// TIA Portal project "uppgift2IndustriellIT" (V18) (continued)
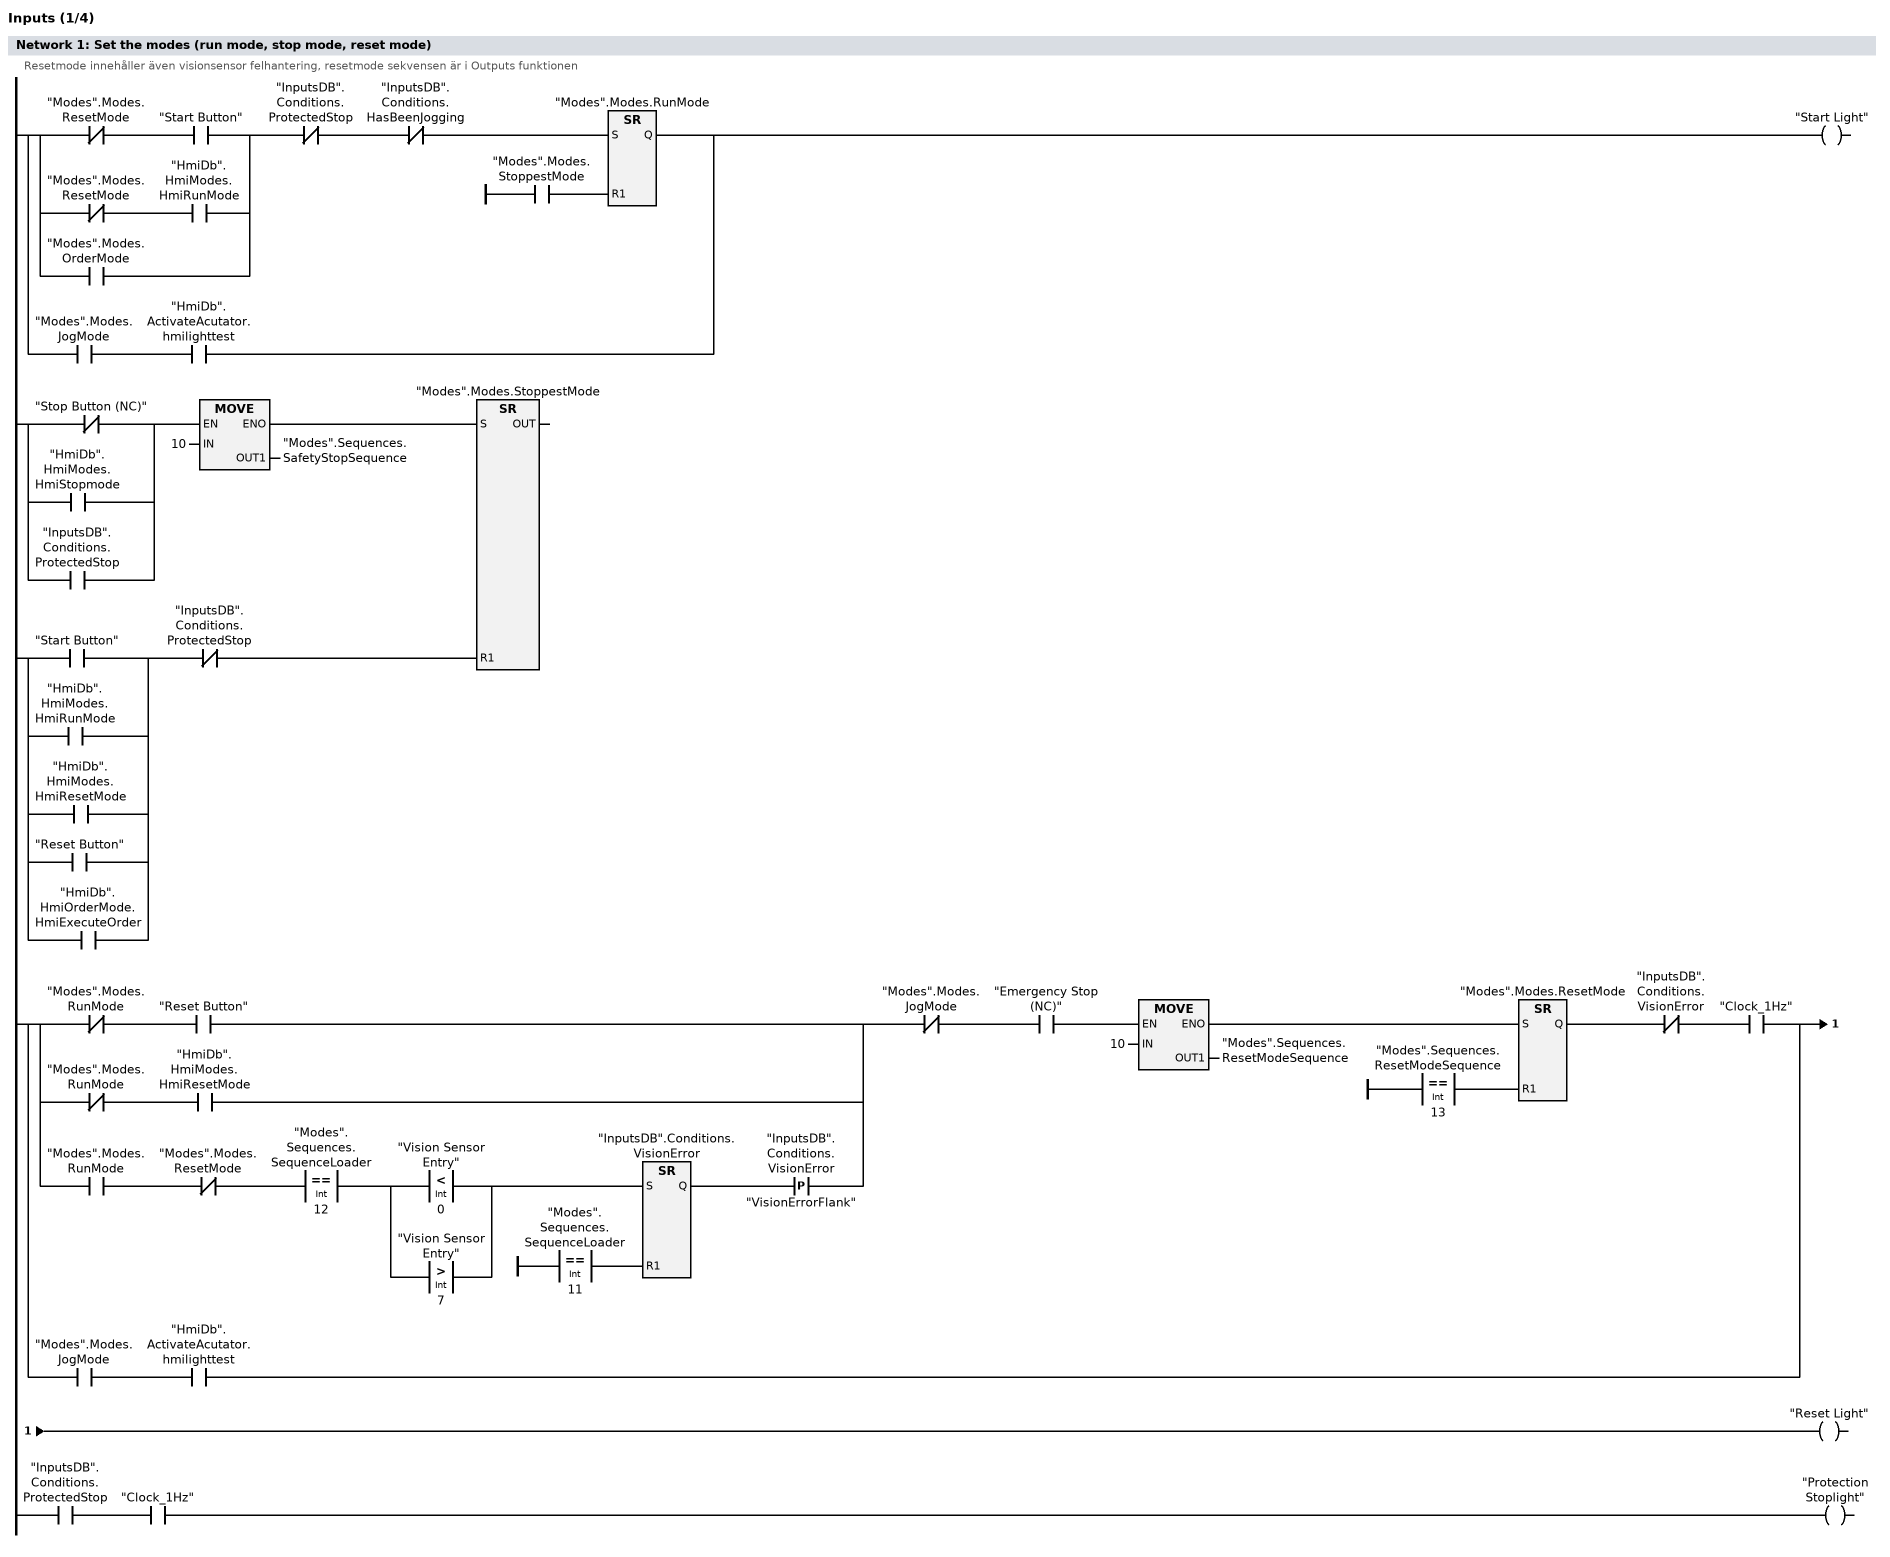
   RUNG wire#powerrail
      I_Contact( "Modes".Modes.ResetMode )
      Contact( "Start Button" )
      wire#w1
      I_Contact( "InputsDB".Conditions.ProtectedStop )
      I_Contact( "InputsDB".Conditions.HasBeenJogging )
      S_SR(operand := "Modes".Modes.RunMode, r1 := wire#w2)
      wire#w3
      Coil( "Start Light" )
   END_RUNG
   RUNG wire#powerrail
      I_Contact( "Modes".Modes.ResetMode )
      Contact( "HmiDb".HmiModes.HmiRunMode )
   END_RUNG wire#w1
   RUNG wire#powerrail
      Contact( "Modes".Modes.OrderMode )
   END_RUNG wire#w1
   RUNG wire#powerrail
      Contact( "Modes".Modes.StoppestMode )
   END_RUNG wire#w2
   RUNG wire#powerrail
      Contact( "Modes".Modes.JogMode )
      Contact( "HmiDb".ActivateAcutator.hmilighttest )
   END_RUNG wire#w3
   RUNG wire#powerrail
      I_Contact( "Stop Button (NC)" )
      wire#w4
      Move(in := 10, out1 => "Modes".Sequences.SafetyStopSequence)
      S_SR(operand := "Modes".Modes.StoppestMode, r1 := wire#w6)
   END_RUNG
   RUNG wire#powerrail
      Contact( "HmiDb".HmiModes.HmiStopmode )
   END_RUNG wire#w4
   RUNG wire#powerrail
      Contact( "InputsDB".Conditions.ProtectedStop )
   END_RUNG wire#w4
   RUNG wire#powerrail
      Contact( "Start Button" )
      wire#w5
      I_Contact( "InputsDB".Conditions.ProtectedStop )
   END_RUNG wire#w6
   RUNG wire#powerrail
      Contact( "HmiDb".HmiModes.HmiRunMode )
   END_RUNG wire#w5
   RUNG wire#powerrail
      Contact( "HmiDb".HmiModes.HmiResetMode )
   END_RUNG wire#w5
   RUNG wire#powerrail
      Contact( "Reset Button" )
   END_RUNG wire#w5
   RUNG wire#powerrail
      Contact( "HmiDb".HmiOrderMode.HmiExecuteOrder )
   END_RUNG wire#w5
   RUNG wire#powerrail
      I_Contact( "Modes".Modes.RunMode )
      Contact( "Reset Button" )
      wire#w7
      I_Contact( "Modes".Modes.JogMode )
      Contact( "Emergency Stop (NC)" )
      Move(in := 10, out1 => "Modes".Sequences.ResetModeSequence)
      S_SR(operand := "Modes".Modes.ResetMode, r1 := wire#w11)
      I_Contact( "InputsDB".Conditions.VisionError )
      Contact( "Clock_1Hz" )
      wire#w12
      Coil( "Reset Light" )
   END_RUNG
   RUNG wire#powerrail
      I_Contact( "Modes".Modes.RunMode )
      Contact( "HmiDb".HmiModes.HmiResetMode )
   END_RUNG wire#w7
   RUNG wire#powerrail
      Contact( "Modes".Modes.RunMode )
      I_Contact( "Modes".Modes.ResetMode )
      { S7_Templates := "SrcType := Int" } EQ_Contact(in1 := "Modes".Sequences.SequenceLoader, in2 := 12)
      wire#w8
      { S7_Templates := "SrcType := Int" } LT_Contact(in1 := "Vision Sensor Entry", in2 := 0)
      wire#w9
      S_SR(operand := "InputsDB".Conditions.VisionError, r1 := wire#w10)
      P_Contact(operand := "InputsDB".Conditions.VisionError, bit := "VisionErrorFlank")
   END_RUNG wire#w7
   RUNG wire#w8
      { S7_Templates := "SrcType := Int" } GT_Contact(in1 := "Vision Sensor Entry", in2 := 7)
   END_RUNG wire#w9
   RUNG wire#powerrail
      { S7_Templates := "SrcType := Int" } EQ_Contact(in1 := "Modes".Sequences.SequenceLoader, in2 := 11)
   END_RUNG wire#w10
   RUNG wire#powerrail
      { S7_Templates := "SrcType := Int" } EQ_Contact(in1 := "Modes".Sequences.ResetModeSequence, in2 := 13)
   END_RUNG wire#w11
   RUNG wire#powerrail
      Contact( "Modes".Modes.JogMode )
      Contact( "HmiDb".ActivateAcutator.hmilighttest )
   END_RUNG wire#w12
   RUNG wire#powerrail
      Contact( "InputsDB".Conditions.ProtectedStop )
      Contact( "Clock_1Hz" )
      Coil( "Protection Stoplight" )
   END_RUNG
   // the same network as SCL:
   IF ((NOT "Modes".Modes.ResetMode AND "Start Button") OR (NOT "Modes".Modes.ResetMode AND "HmiDb".HmiModes.HmiRunMode) OR "Modes".Modes.OrderMode) AND NOT "InputsDB".Conditions.ProtectedStop AND NOT "InputsDB".Conditions.HasBeenJogging THEN
       "Modes".Modes.RunMode := TRUE;   // SR flip-flop
   END_IF;
   IF "Modes".Modes.StoppestMode THEN "Modes".Modes.RunMode := FALSE; END_IF;
   "Start Light" := "Modes".Modes.RunMode OR ("Modes".Modes.JogMode AND "HmiDb".ActivateAcutator.hmilighttest);
   #_w1 := NOT "Stop Button (NC)" OR "HmiDb".HmiModes.HmiStopmode OR "InputsDB".Conditions.ProtectedStop;
   IF #_w1 THEN
       "Modes".Sequences.SafetyStopSequence := 10;
       "Modes".Modes.StoppestMode := TRUE;   // SR flip-flop
   END_IF;
   IF ("Start Button" OR "HmiDb".HmiModes.HmiRunMode OR "HmiDb".HmiModes.HmiResetMode OR "Reset Button" OR "HmiDb".HmiOrderMode.HmiExecuteOrder) AND NOT "InputsDB".Conditions.ProtectedStop THEN
       "Modes".Modes.StoppestMode := FALSE;
   END_IF;
   IF "Modes".Modes.RunMode AND NOT "Modes".Modes.ResetMode AND ("Modes".Sequences.SequenceLoader = 12) AND (("Vision Sensor Entry" < 0) OR ("Vision Sensor Entry" > 7)) THEN
       "InputsDB".Conditions.VisionError := TRUE;   // SR flip-flop
   END_IF;
   IF "Modes".Sequences.SequenceLoader = 11 THEN "InputsDB".Conditions.VisionError := FALSE; END_IF;
   #_w2 := "InputsDB".Conditions.VisionError AND "InputsDB".Conditions.VisionError AND NOT "VisionErrorFlank";   // rising edge of "InputsDB".Conditions.VisionError
   "VisionErrorFlank" := "InputsDB".Conditions.VisionError;
   #_w3 := ((NOT "Modes".Modes.RunMode AND "Reset Button") OR (NOT "Modes".Modes.RunMode AND "HmiDb".HmiModes.HmiResetMode) OR #_w2) AND NOT "Modes".Modes.JogMode AND "Emergency Stop (NC)";
   IF #_w3 THEN
       "Modes".Sequences.ResetModeSequence := 10;
       "Modes".Modes.ResetMode := TRUE;   // SR flip-flop
   END_IF;
   IF "Modes".Sequences.ResetModeSequence = 13 THEN "Modes".Modes.ResetMode := FALSE; END_IF;
   "Reset Light" := ("Modes".Modes.ResetMode AND NOT "InputsDB".Conditions.VisionError AND "Clock_1Hz") OR ("Modes".Modes.JogMode AND "HmiDb".ActivateAcutator.hmilighttest);
   "Protection Stoplight" := "InputsDB".Conditions.ProtectedStop AND "Clock_1Hz";
END_REGION

REGION Network 2: Activate Stop light
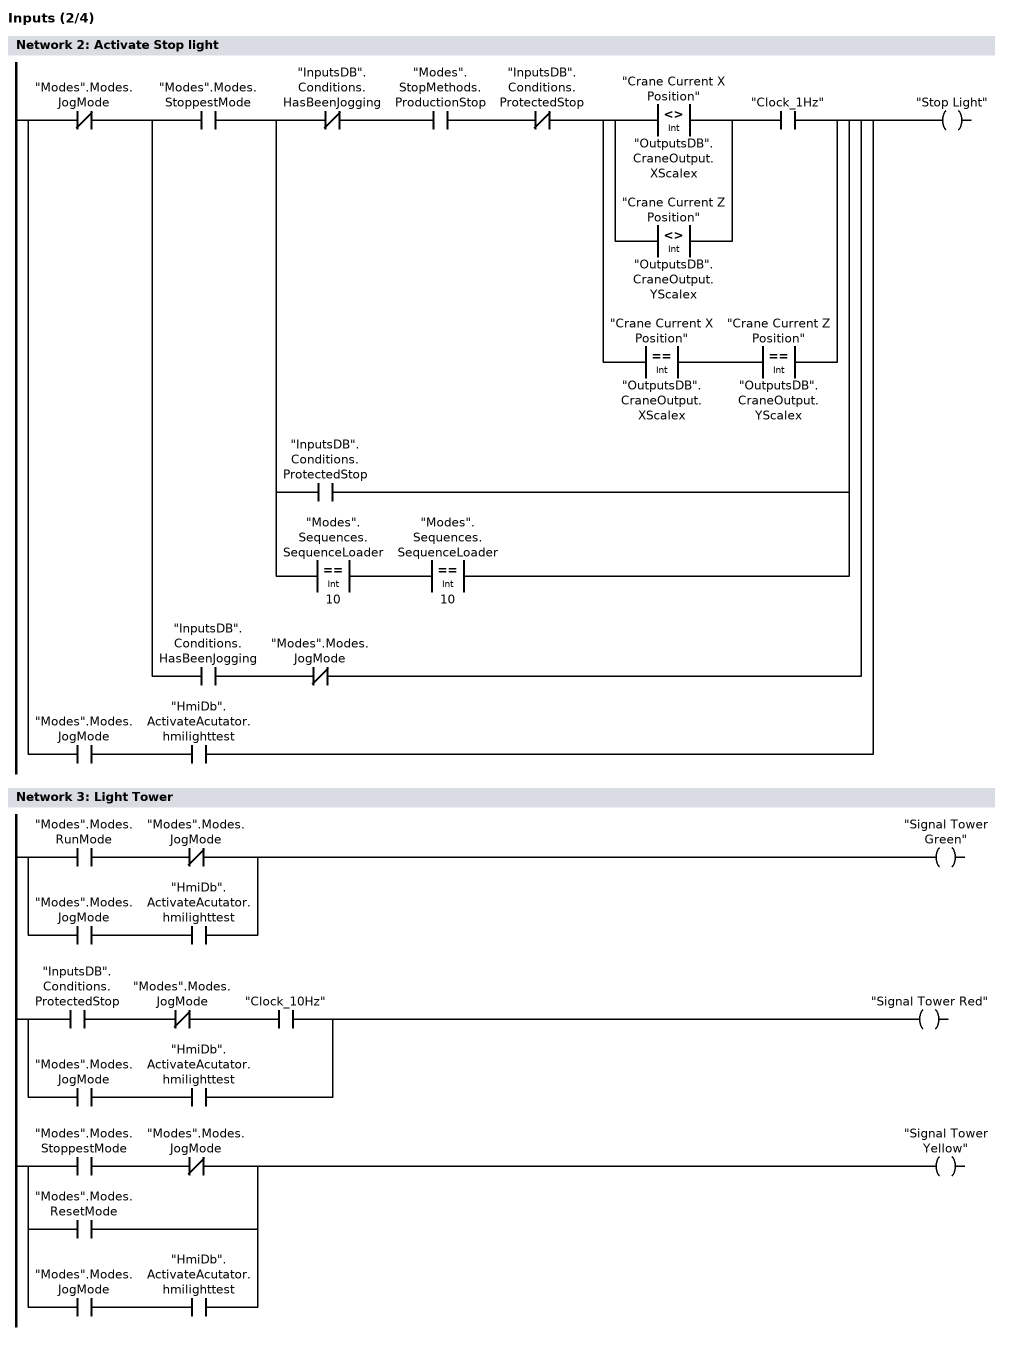
   RUNG wire#powerrail
      I_Contact( "Modes".Modes.JogMode )
      wire#w1
      Contact( "Modes".Modes.StoppestMode )
      wire#w2
      I_Contact( "InputsDB".Conditions.HasBeenJogging )
      Contact( "Modes".StopMethods.ProductionStop )
      I_Contact( "InputsDB".Conditions.ProtectedStop )
      wire#w3
      { S7_Templates := "SrcType := Int" } NE_Contact(in1 := "Crane Current X Position", in2 := "OutputsDB".CraneOutput.XScalex)
      wire#w4
      Contact( "Clock_1Hz" )
      wire#w5
      Coil( "Stop Light" )
   END_RUNG
   RUNG wire#w3
      { S7_Templates := "SrcType := Int" } NE_Contact(in1 := "Crane Current Z Position", in2 := "OutputsDB".CraneOutput.YScalex)
   END_RUNG wire#w4
   RUNG wire#w3
      { S7_Templates := "SrcType := Int" } EQ_Contact(in1 := "Crane Current X Position", in2 := "OutputsDB".CraneOutput.XScalex)
      { S7_Templates := "SrcType := Int" } EQ_Contact(in1 := "Crane Current Z Position", in2 := "OutputsDB".CraneOutput.YScalex)
   END_RUNG wire#w5
   RUNG wire#w2
      Contact( "InputsDB".Conditions.ProtectedStop )
   END_RUNG wire#w5
   RUNG wire#w2
      { S7_Templates := "SrcType := Int" } EQ_Contact(in1 := "Modes".Sequences.SequenceLoader, in2 := 10)
      { S7_Templates := "SrcType := Int" } EQ_Contact(in1 := "Modes".Sequences.SequenceLoader, in2 := 10)
   END_RUNG wire#w5
   RUNG wire#w1
      Contact( "InputsDB".Conditions.HasBeenJogging )
      I_Contact( "Modes".Modes.JogMode )
   END_RUNG wire#w5
   RUNG wire#powerrail
      Contact( "Modes".Modes.JogMode )
      Contact( "HmiDb".ActivateAcutator.hmilighttest )
   END_RUNG wire#w5
   // the same network as SCL:
   "Stop Light" := (NOT "Modes".Modes.JogMode AND (("Modes".Modes.StoppestMode AND ((NOT "InputsDB".Conditions.HasBeenJogging AND "Modes".StopMethods.ProductionStop AND NOT "InputsDB".Conditions.ProtectedStop AND (((("Crane Current X Position" <> "OutputsDB".CraneOutput.XScalex) OR ("Crane Current Z Position" <> "OutputsDB".CraneOutput.YScalex)) AND "Clock_1Hz") OR (("Crane Current X Position" = "OutputsDB".CraneOutput.XScalex) AND ("Crane Current Z Position" = "OutputsDB".CraneOutput.YScalex)))) OR "InputsDB".Conditions.ProtectedStop OR (("Modes".Sequences.SequenceLoader = 10) AND ("Modes".Sequences.SequenceLoader = 10)))) OR ("InputsDB".Conditions.HasBeenJogging AND NOT "Modes".Modes.JogMode))) OR ("Modes".Modes.JogMode AND "HmiDb".ActivateAcutator.hmilighttest);
END_REGION

REGION Network 3: Light Tower
   RUNG wire#powerrail
      Contact( "Modes".Modes.RunMode )
      I_Contact( "Modes".Modes.JogMode )
      wire#w1
      Coil( "Signal Tower Green" )
   END_RUNG
   RUNG wire#powerrail
      Contact( "Modes".Modes.JogMode )
      Contact( "HmiDb".ActivateAcutator.hmilighttest )
   END_RUNG wire#w1
   RUNG wire#powerrail
      Contact( "InputsDB".Conditions.ProtectedStop )
      I_Contact( "Modes".Modes.JogMode )
      Contact( "Clock_10Hz" )
      wire#w2
      Coil( "Signal Tower Red" )
   END_RUNG
   RUNG wire#powerrail
      Contact( "Modes".Modes.JogMode )
      Contact( "HmiDb".ActivateAcutator.hmilighttest )
   END_RUNG wire#w2
   RUNG wire#powerrail
      Contact( "Modes".Modes.StoppestMode )
      I_Contact( "Modes".Modes.JogMode )
      wire#w3
      Coil( "Signal Tower Yellow" )
   END_RUNG
   RUNG wire#powerrail
      Contact( "Modes".Modes.ResetMode )
   END_RUNG wire#w3
   RUNG wire#powerrail
      Contact( "Modes".Modes.JogMode )
      Contact( "HmiDb".ActivateAcutator.hmilighttest )
   END_RUNG wire#w3
   // the same network as SCL:
   "Signal Tower Green" := ("Modes".Modes.RunMode AND NOT "Modes".Modes.JogMode) OR ("Modes".Modes.JogMode AND "HmiDb".ActivateAcutator.hmilighttest);
   "Signal Tower Red" := ("InputsDB".Conditions.ProtectedStop AND NOT "Modes".Modes.JogMode AND "Clock_10Hz") OR ("Modes".Modes.JogMode AND "HmiDb".ActivateAcutator.hmilighttest);
   "Signal Tower Yellow" := ("Modes".Modes.StoppestMode AND NOT "Modes".Modes.JogMode) OR "Modes".Modes.ResetMode OR ("Modes".Modes.JogMode AND "HmiDb".ActivateAcutator.hmilighttest);
END_REGION

REGION Network 4: Crane raw sensor value to MM
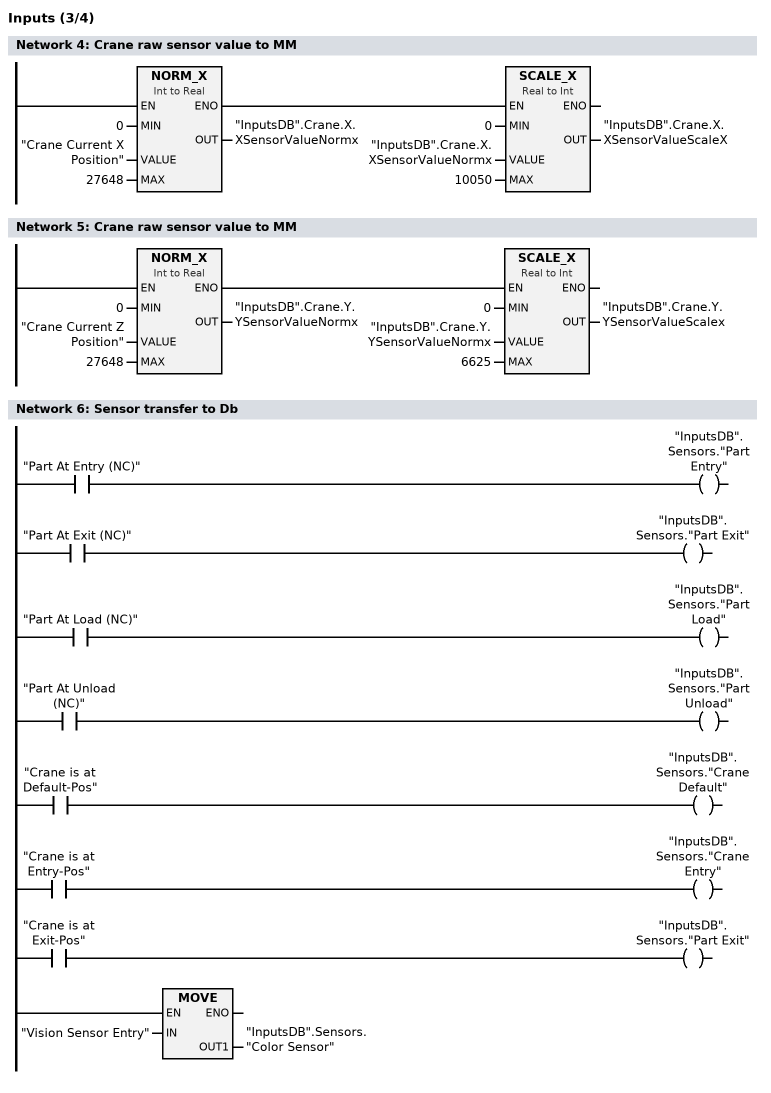
   RUNG wire#powerrail
      { S7_Templates := "[SrcType := Int, DestType := Real]" } Normalize(min := 0, value := "Crane Current X Position", max := 27648, out => "InputsDB".Crane.X.XSensorValueNormx)
      { S7_Templates := "[SrcType := Real, DestType := Int]" } Scale(min := 0, value := "InputsDB".Crane.X.XSensorValueNormx, max := 10050, out => "InputsDB".Crane.X.XSensorValueScaleX)
   END_RUNG
   // the same network as SCL:
   "InputsDB".Crane.X.XSensorValueNormx := NORM_X(MIN := 0, VALUE := "Crane Current X Position", MAX := 27648);
   "InputsDB".Crane.X.XSensorValueScaleX := SCALE_X(MIN := 0, VALUE := "InputsDB".Crane.X.XSensorValueNormx, MAX := 10050);
END_REGION

REGION Network 5: Crane raw sensor value to MM
   RUNG wire#powerrail
      { S7_Templates := "[SrcType := Int, DestType := Real]" } Normalize(min := 0, value := "Crane Current Z Position", max := 27648, out => "InputsDB".Crane.Y.YSensorValueNormx)
      { S7_Templates := "[SrcType := Real, DestType := Int]" } Scale(min := 0, value := "InputsDB".Crane.Y.YSensorValueNormx, max := 6625, out => "InputsDB".Crane.Y.YSensorValueScalex)
   END_RUNG
   // the same network as SCL:
   "InputsDB".Crane.Y.YSensorValueNormx := NORM_X(MIN := 0, VALUE := "Crane Current Z Position", MAX := 27648);
   "InputsDB".Crane.Y.YSensorValueScalex := SCALE_X(MIN := 0, VALUE := "InputsDB".Crane.Y.YSensorValueNormx, MAX := 6625);
END_REGION

REGION Network 6: Sensor transfer to Db
   RUNG wire#powerrail
      Contact( "Part At Entry (NC)" )
      Coil( "InputsDB".Sensors."Part Entry" )
   END_RUNG
   RUNG wire#powerrail
      Contact( "Part At Exit (NC)" )
      Coil( "InputsDB".Sensors."Part Exit" )
   END_RUNG
   RUNG wire#powerrail
      Contact( "Part At Load (NC)" )
      Coil( "InputsDB".Sensors."Part Load" )
   END_RUNG
   RUNG wire#powerrail
      Contact( "Part At Unload (NC)" )
      Coil( "InputsDB".Sensors."Part Unload" )
   END_RUNG
   RUNG wire#powerrail
      Contact( "Crane is at Default-Pos" )
      Coil( "InputsDB".Sensors."Crane Default" )
   END_RUNG
   RUNG wire#powerrail
      Contact( "Crane is at Entry-Pos" )
      Coil( "InputsDB".Sensors."Crane Entry" )
   END_RUNG
   RUNG wire#powerrail
      Contact( "Crane is at Exit-Pos" )
      Coil( "InputsDB".Sensors."Part Exit" )
   END_RUNG
   RUNG wire#powerrail
      Move(in := "Vision Sensor Entry", out1 => "InputsDB".Sensors."Color Sensor")
   END_RUNG
   // the same network as SCL:
   "InputsDB".Sensors."Part Entry" := "Part At Entry (NC)";
   "InputsDB".Sensors."Part Exit" := "Part At Exit (NC)";
   "InputsDB".Sensors."Part Load" := "Part At Load (NC)";
   "InputsDB".Sensors."Part Unload" := "Part At Unload (NC)";
   "InputsDB".Sensors."Crane Default" := "Crane is at Default-Pos";
   "InputsDB".Sensors."Crane Entry" := "Crane is at Entry-Pos";
   "InputsDB".Sensors."Part Exit" := "Crane is at Exit-Pos";
   "InputsDB".Sensors."Color Sensor" := "Vision Sensor Entry";
END_REGION

REGION Network 7: counter free slots
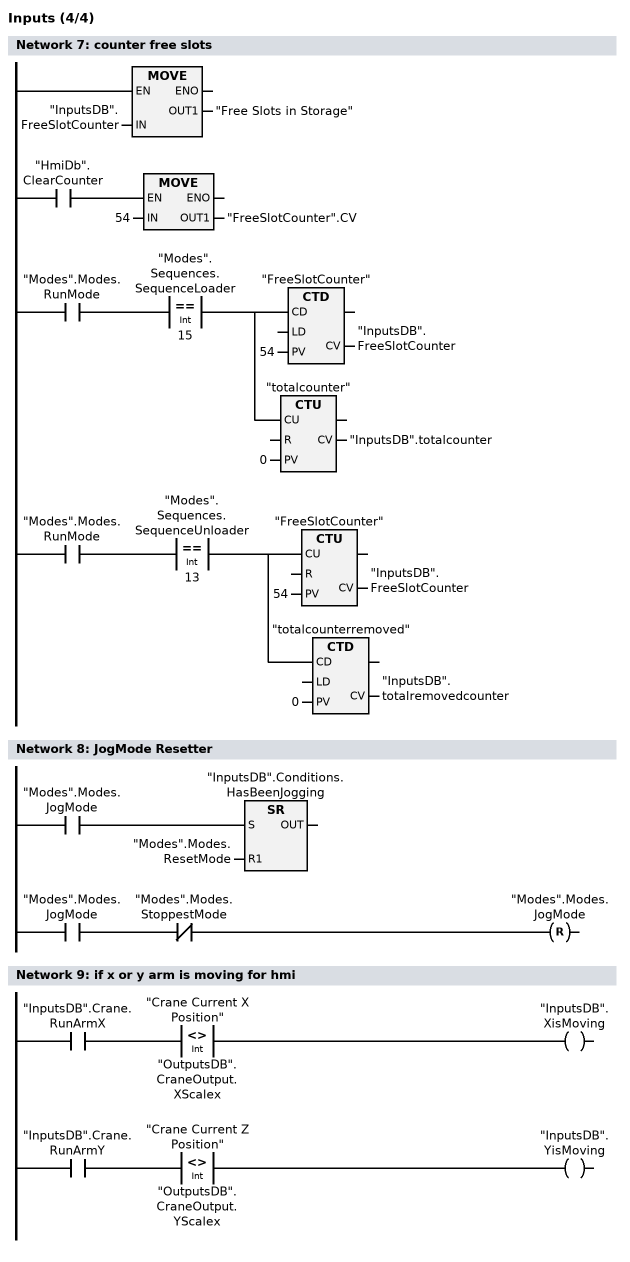
   "Free Slots in Storage" := "InputsDB".FreeSlotCounter;
   IF "HmiDb".ClearCounter THEN "FreeSlotCounter".CV := 54; END_IF;
   #_w1 := "Modes".Modes.RunMode AND ("Modes".Sequences.SequenceLoader = 15);
   "FreeSlotCounter".CTD(CD := #_w1, PV := 54, CV => "InputsDB".FreeSlotCounter);
   "totalcounter".CTU(CU := #_w1, PV := 0, CV => "InputsDB".totalcounter);
   #_w2 := "Modes".Modes.RunMode AND ("Modes".Sequences.SequenceUnloader = 13);
   "FreeSlotCounter".CTU(CU := #_w2, PV := 54, CV => "InputsDB".FreeSlotCounter);
   "totalcounterremoved".CTD(CD := #_w2, PV := 0, CV => "InputsDB".totalremovedcounter);
END_REGION

REGION Network 8: JogMode Resetter
   RUNG wire#powerrail
      Contact( "Modes".Modes.JogMode )
      S_SR(operand := "InputsDB".Conditions.HasBeenJogging, r1 := "Modes".Modes.ResetMode)
   END_RUNG
   RUNG wire#powerrail
      Contact( "Modes".Modes.JogMode )
      I_Contact( "Modes".Modes.StoppestMode )
      R_Coil( "Modes".Modes.JogMode )
   END_RUNG
   // the same network as SCL:
   IF "Modes".Modes.JogMode THEN
       "InputsDB".Conditions.HasBeenJogging := TRUE;   // SR flip-flop
   END_IF;
   IF "Modes".Modes.ResetMode THEN "InputsDB".Conditions.HasBeenJogging := FALSE; END_IF;
   IF "Modes".Modes.JogMode AND NOT "Modes".Modes.StoppestMode THEN "Modes".Modes.JogMode := FALSE; END_IF;
END_REGION
